// TIA Portal project "E95238_MCC1200_Sisecam_India" (V17) (continued)
TYPE "UDT_CapData_Tracking"
   STRUCT
      dTrackingHead : DInt;   // Tracking head on the circular buffer
      dTrackingTail : DInt;   // Tracking tail on the circular buffer
      dLastInsertIndex : DInt;   // Last insert index on circular
      dLastTargetLineValue_cmm : DInt;   // Last target line value [mm/100]
      dNextValidCapID : DInt;   // Next valid cap ID
      dLastValidCapID : DInt;   // Last valid cap ID
      dMutexCounter : DInt;   // Mutex counter for thread safe
      xInsertCapOnTrack : Bool;   // Insert cap on tracking
      timeLastAccessMutex : Time;   // Time of the last access mutex
      rgxNewCapAvailable : Array[0.."DMAXELEMWAKEUPNEWPLATE_IND"] of Bool;   // New cap available for other machines. Machines not used should be manually resetted
      tNewCapToInsert : "UDT_CapData";   // New cap to insert on tracking
      tLastPlacedCap : "UDT_CapData";   // Last placed cap on tracking
      rgtTrackCaps : Array[0.."DMAXTRACKCAP_IND"] of Struct   // Buffer of caps
         dEncValueHeadSnaproll_cmm : DInt;   // Encoder value on snap roll head [mm/100]
         dEncValueTailSnaproll_cmm : DInt;   // Encoder value on snap roll tail [mm/100]
         tCap : "UDT_CapData";   // Cap data
         rgxMachineExecMask : Array[0.."DMAXTRACKMACHINE_IND"] of Bool;   // Machine execution mask
      END_STRUCT;
      rgtTrackMachine : Array[0.."DMAXTRACKMACHINE_IND"] of Struct   // Tracking machine
         tUserData : Struct   // User data
            dSetDistanceSnap_cmm : DInt;   // Distance from snaproll [mm/100]
            dSetMachReacTime_ms : DInt;   // Machine reaction time [ms] (Positive to anticipate / Negative to delay)
            xGetPosReach : Bool;   // New cap arrive on position
            dGetUpstremIndex : DInt;   // Upstream cap position index
            dGetDownstreamIndex : DInt;   // Downstream cap position index
            dGetEncValueOnSnap_cmm : DInt;   // Encoder value on snaproll [mm/100]
         END_STRUCT;
         tAuxData : Struct   // Internal data for tracking
            dActualMachineEncValue_cmm : DInt;   // Actual machine encoder value [mm/100]
            dPrevCapIndex : DInt;   // Previous cap index
            dNextCapIndex : DInt;   // Next cap index
         END_STRUCT;
      END_STRUCT;
      tEmptyCap : "UDT_CapData";   // Cap with empty data (used for initialization)
      rgtTrackSearch : Array[0.."DMAXELEMTRACKSEARCH_IND"] of Struct   // Tracking search data
         xRequestSearchPlate : Bool;   // Request search plate
         xPlateFound : Bool;   // Plate found by tracking
         dRequestID : DInt;   // Number to identify the request
         dAnalyzedID : DInt;   // Number to identify the processed request
         dFoundTrackIndex : DInt;   // Plate pointer ID founded
         dSearchMode : DInt;   // Search mode (1=Limit head, 2=Limit tail 3=Both)
         dMinHeadPosition_cmm : DInt;   // Minimum head position distance from snaproll [mm/100]
         dMaxHeadPosition_cmm : DInt;   // Maximum head position distance from snaproll [mm/100]
         dMinTailPosition_cmm : DInt;   // Minumum tail position distance from snaproll [mm/100]
         dMaxTailPosition_cmm : DInt;   // Maximum tail position distance from snaproll [mm/100]
         tSearchRequest : Struct   // Search request
            xMainDestEqual : Bool;   // Main destination equal
            xLengthLessThan : Bool;   // Cap length is less than
            xCutDone : Bool;   // XCut is done
            xSpare_3 : Bool;
            xSpare_4 : Bool;
            xSpare_5 : Bool;
            xSpare_6 : Bool;
            xSpare_7 : Bool;
            xSpare_8 : Bool;
            xSpare_9 : Bool;
            xSpare_10 : Bool;
            xSpare_11 : Bool;
            xSpare_12 : Bool;
            xSpare_13 : Bool;
            xSpare_14 : Bool;
            xSpare_15 : Bool;
            xSpare_16 : Bool;
            xSpare_17 : Bool;
            xSpare_18 : Bool;
            xSpare_19 : Bool;
            xSpare_20 : Bool;
            xSpare_21 : Bool;
            xSpare_22 : Bool;
            xSpare_23 : Bool;
            xSpare_24 : Bool;
            xSpare_25 : Bool;
            xSpare_26 : Bool;
            xSpare_27 : Bool;
            xSpare_28 : Bool;
            xSpare_29 : Bool;
            xSpare_30 : Bool;
            xSpare_31 : Bool;
         END_STRUCT;
         tSearchData : Struct
            dMainDest_mask : LInt;   // Main destination mask
            dLength_cmm : DInt;   // Length [mm/100]
         END_STRUCT;
      END_STRUCT;
   END_STRUCT;
END_TYPE

// folder: 03_Encoder

TYPE "UDT_Encoder"
   STRUCT
      dActualEncoderCounter_cmm : DInt;   // Actual encoder counter [mm/100]
      rActSpeedValue_cmm_ms : Real;   // Actual speed value [(mm/100)/ms]
      dActSpeedValue_mm_min : DInt;   // Actual speed value [mm/min]
      rActSpeedValueFast_cmm_ms : Real;   // Actual speed value updated 500ms [(mm/100)/ms]
      dActSpeedValueFast_mm_min : DInt;   // Actual speed value updated 500ms [mm/min]
      dLastMeterValue_cmm : DInt;   // Last meter counter value [mm/100]
      dNextMeterValue_cmm : DInt;   // Next meter counter value [mm/100]
      rgxMetersForXcuts : Array[0.."DMAXXHEADS_IND"] of Bool;   // Meters signal for XCuts
      rgxMetersForYCuts : Array[0.."DMAXYCUTBRIDGE_IND"] of Bool;   // Meters signal for YCuts
      xMeterForMarkers : Bool;   // Meter signal for Markers
      xMeterForScanner : Bool;   // Meter signal for Scanner
   END_STRUCT;
END_TYPE

TYPE "LPD_typeCountFeedbackCh"
VERSION : 0.1
   STRUCT
      countValue : DInt := 16#0000;   // Current count value
      capturedValue : DInt := 16#0000;   // Last Capture value acquired
      measuredValue : Real := 0.0;   // Current measured value
      powerError : Bool := FALSE;   // Incorrect supply voltage L+
      encError : Bool := FALSE;   // Incorrect encoder signal
      ldError : Bool := FALSE;   // Error when loading via control interface
      reserved1 : Bool := FALSE;   // Reserved
      reserved2 : Bool := FALSE;   // Reserved
      reserved3 : Bool := FALSE;   // Reserved
      reserved4 : Bool := FALSE;   // Reserved
      reserved5 : Bool := FALSE;   // Reserved
      commActive : Bool := FALSE;   // Comm active
      resEventAck : Bool := FALSE;   // Reset of event bits active
      ldStsSlot0 : Bool := FALSE;   // Load request for Slot 0 detected and executed (toggling)
      ldStsSlot1 : Bool := FALSE;   // Load request for Slot 1 detected and executed (toggling)
      stsReady : Bool := FALSE;   // Digital on-board I/O started up and parameters assigned
      stsSwGate : Bool := FALSE;   // Software gate status
      reserved7 : Bool := FALSE;   // Reserved
      reserved8 : Bool := FALSE;   // Reserved
      stsDir : Bool := FALSE;   // Direction of last count value change
      stsCount : Bool := FALSE;   // Count pulse detected within last approx. 0.5 s
      stsGate : Bool := FALSE;   // Internal gate status
      stsDQ0 : Bool := FALSE;   // Status HSC DQ0
      stsDQ1 : Bool := FALSE;   // Status HSC DQ1
      stsDI0 : Bool := FALSE;   // Status HSC DI0
      stsDI1 : Bool := FALSE;   // Status HSC DI1
      stsDI2 : Bool := FALSE;   // Status HSC DI2
      eventZero : Bool := FALSE;   // Zero crossing has occurred
      eventUnderflow : Bool := FALSE;   // Underflow has occurred
      eventOverflow : Bool := FALSE;   // Overflow has occurred
      eventCompare0 : Bool := FALSE;   // Comparison event for DQ0 has occurred
      eventCompare1 : Bool := FALSE;   // Comparison event for DQ1 has occurred
      eventSync : Bool := FALSE;   // Synchronization has occurred
      eventCapture : Bool := FALSE;   // Capture event has occurred
      stsMeasInterval : Bool := FALSE;   // Count pulse detected in previous measuring interval
   END_STRUCT;
END_TYPE

TYPE "LPD_typeCountControlCh"
VERSION : 0.1
   STRUCT
      loadValue0 : DWord := 16#0000;   // Load value 0
      loadValue1 : DWord := 16#0000;   // Load value 1
      controlByte : Byte := B#16#00;   // Control byte load value
      swGate : Bool := FALSE;   // Software gate
      tmCtrlDQ0 : Bool := FALSE;   // Enable technological function DQ0
      tmCtrlDQ1 : Bool := FALSE;   // Enable technological function DQ1
      setDQ0 : Bool := FALSE;   // Set DQ0
      setDQ1 : Bool := FALSE;   // Set DQ1
      enSyncUp : Bool := FALSE;   // Enable upward synchronization
      enSyncDown : Bool := FALSE;   // Enable downward synchronization
      enCapture : Bool := FALSE;   // Enable capture function
      resError : Bool := FALSE;   // Reset of saved error states
      resEvent : Bool := FALSE;   // Reset of saved events
      reserved0 : Bool := FALSE;   // Reserved
      reserved1 : Bool := FALSE;   // Reserved
      reserved2 : Bool := FALSE;   // Reserved
      reserved3 : Bool := FALSE;   // Reserved
      reserved4 : Bool := FALSE;   // Reserved
      SetDir : Bool := FALSE;   // Count direction (with encoder without direction signal)
      reserved5 : Byte;   // Reserved
   END_STRUCT;
END_TYPE

// folder: 04_XCuts

TYPE "UDT_XCUT_DRIVE_INPUT"
   STRUCT
      rgxStatusBits : Struct
         xFault_EmergencyON : Bool := false;   // DN_SMAPP_FEMERGENCY_ON
         xFault_AuxPowerOFF : Bool := false;   // DN_SMAPP_FAUXPOWER_OFF
         xFault_InputPowerOFF : Bool := false;   // DN_SMAPP_FINPPOWER_OFF
         xFault_SafetyArea : Bool := false;   // DN_SMAPP_FSAFETYAREA
         xFault_Overtstroke : Bool := false;   // DN_SMAPP_FOVERSTROKE
         xFaultl_OverTemp : Bool := false;   // DN_SMAPP_FOVERTEMP
         xFault_CarriageNotDown : Bool := false;   // DN_SMAPP_FCARRIAGEDOWN
         xFault_MissingAir : Bool := false;   // DN_SMAPP_FMISSINGAIR
         xFault_AxisFault : Bool := false;   // DN_SMAPP_FAXISFAULT
         xFault_DriveNotEnable : Bool := false;   // DN_SMAPP_FDRIVENOENABLE
         xFault_TankOilEmpty : Bool := false;   // DN_SMAPP_FTANKOILEMPTY
         xFault_CarriageOff : Bool := false;   // DN_SMAPP_FCARRIAGEOFF
         xFault_ExtInpPower : Bool := false;   // DN_SMAPP_FEXTINPPOWER
         xFault_EmergencyLoc1 : Bool := false;   // DN_SMAPP_FLOCALEMERG_1
         xFault_EmergencyLoc2 : Bool := false;   // DN_SMAPP_FLOCALEMERG_2
         xFault_EmergencyLoc3 : Bool := false;   // DN_SMAPP_FLOCALEMERG_3
         xStatus_AxisOnline : Bool := false;   // DN_SMAPP_AXISONLINE
         xStatus_AxisReady : Bool := false;   // DN_SMAPP_AXISREADY
         xStatus_HomeProgress : Bool := false;   // DN_SMAPP_HOMEPROGRESS
         xStatus_MoveProgress : Bool := false;   // DN_SMAPP_MOVEPROGRESS
         xStatus_MoveProgrNick : Bool := false;   // DN_SMAPP_MOVEPROGRESSNICK
         xStatus_InvertReady : Bool := false;   // DN_SMAPP_INVERTERREADY
         xStatus_BridgeEnabled : Bool := false;   // DN_SMAPP_BRIDGEENABLED
         xStatus_AxisSyncronized : Bool := false;   // DN_SMAPP_AXISSYNCRONIZED
         xStatus_ButtonEnabled : Bool;   // Button enabled
         xStatus_xSpare17 : Bool;   // Spare
         xStatus_xSpare18 : Bool;   // Spare
         xStatus_xSpare19 : Bool;   // Spare
         xStatus_xSpare20 : Bool;   // Spare
         xStatus_xSpare21 : Bool;   // Spare
         xStatus_xSpare22 : Bool;   // Spare
         xStatus_xSpare23 : Bool;   // Spare
      END_STRUCT;
      dCarriagePos_dmm : DInt := 0;   // DN_SMAPP_CARRIAGEPOS [mm/10]
      dLehrPosition_cmm : DInt := 0;   // DN_SMAPP_LEHRPOSITION [mm/100]
      dLehrSpeed_cmm_min : DInt := 0;   // DN_SMAPP_LEHRSPEED [mm/10/min]
      dErrorCode : DInt := 0;   // DN_SMAPP_ERRORCODE
      dMissionDone : DInt := 0;   // DN_SMAPP_MISSIONDONE
      dMissionUnDone : DInt := 0;   // DN_SMAPP_MISSION_UNDONE
      iLiveCounter : Int := 0;   // DN_SMAPP_LIVECOUNTER
      iTimeHeadDown_ms : Int;   // Time head down% [ms]
   END_STRUCT;
END_TYPE

TYPE "UDT_XCUT_DRIVE_OUTPUT"
   STRUCT
      rgxControlBits : Struct
         xSpare0 : Bool;
         xSpare1 : Bool;
         xSpare2 : Bool;
         xSpare3 : Bool;
         xFaultReset : Bool := false;   // DN_PLC_FAULTRESET
         xEnableBridge : Bool := false;   // DN_PLC_ENABLEBRIDGE
         xDisableBridge : Bool := false;   // DN_PLC_DISABLEBRIDGE
         xSimulationMode : Bool := false;   // DN_PLC_SIMULATIONMODE
         xDisableRequest : Bool;   // DN_PLC_DISABLEREQUEST
         xSpare9 : Bool;
         xSpare10 : Bool;
         xSpare11 : Bool;
         xSpare12 : Bool;
         xSpare13 : Bool;
         xSpare14 : Bool;
         xSpare15 : Bool;
         xSpare16 : Bool;
         xSpare17 : Bool;
         xSpare18 : Bool;
         xSpare19 : Bool;
         xSpare20 : Bool := false;
         xSpare21 : Bool := false;
         xSpare22 : Bool := false;
         xSpare23 : Bool := false;
         xSpare24 : Bool;
         xSpare25 : Bool;
         xSpare26 : Bool;
         xSpare27 : Bool;
         xSpare28 : Bool;
         xSpare29 : Bool;
         xSpare30 : Bool;
         xSpare31 : Bool;
      END_STRUCT;
      dBridgeAngle_degre_10000 : DInt := 0;   // DN_PLC_BRIDGEANGLE
      dHeadDownPos_dmm : DInt := 0;   // DN_PLC_HEADDOWNPOS
      dHeadRisePos_dmm : DInt := 0;   // DN_PLC_HEADRISEPOS
      iReturnSpeed_rpm : Int := 0;   // DN_PLC_RETURNSPEED
      iTimeHeadDown_ms : Int := 0;   // DN_PLC_TIMEHEADDOWN
      iTimeHeadUp_ms : Int := 0;   // DN_PLC_TIMEHEADUP
      iLubAdvanceTime_ms : Int := 0;   // DN_PLC_LUBADVANCETIME
      iLubDelayTime_ms : Int := 0;   // DN_PLC_LUBDELAYTIME
      iTimeHeadAct_ms : Int := 0;   // DN_PLC_TIMEHEADACTIV
      iTimeHeadDeactiv_ms : Int := 0;   // DN_PLC_TIMEHEADDEACTIV
      dPressure_mN : DInt := 0;   // DN_PLC_PRESSURE
      dMissionID : DInt := 0;   // DN_PLC_MISSIONID
      dMissionCounter : DInt := 0;   // DN_PLC_MISSIONCOUNTER
      dSyncroCounter : DInt := 0;   // DN_PLC_SYNCROCOUNTER
      iLiveCounter : Int := 0;   // DN_PLC_LIVECOUNTER
   END_STRUCT;
END_TYPE

TYPE "UDT_XCUT_AXIS_REF"
   STRUCT
      udi_ModbusAddress_read : UDInt;
      di_ParameterReadValue : DInt;
      x_CommandReadParameter : Bool;
      x_StatusReadParameter_OK : Bool;
      x_StatusReadParameter_Error : Bool;
      udi_ModbusAddress_write : UDInt;
      di_ParameterWriteValue : DInt;
      x_CommandWriteParameter : Bool;
      x_Status_WriteParameter_OK : Bool;
      x_Status_WriteParameter_Error : Bool;
   END_STRUCT;
END_TYPE

// folder: 05_YCuts

TYPE "UDT_YCut_IdeviceToBridge"
   STRUCT
      dSpare1 : Array[0..2] of DInt;
      xCycleON : Bool;
      xResetAnomaly : Bool;
      xResetBuffers : Bool;
      xGlassBreak : Bool;
      xPLCActive0 : Bool;
      xPLCActive1 : Bool;
      xQLTplate : Bool;
      xSpare2 : Bool;
      xSpare3 : Bool;
      xSpare4 : Bool;
      xSpare5 : Bool;
      xSpare6 : Bool;
      xSpare7 : Bool;
      xSpare8 : Bool;
      xSpare9 : Bool;
      xSpare10 : Bool;
      xStatusSpare : Array[0..15] of Bool;
      dSpare2 : Array[0..7] of DInt;
      iSpare : Int;
   END_STRUCT;
END_TYPE

TYPE "UDT_YCut_IdeviceFromBridge"
   STRUCT
      dProcessingIDPlate : DInt;   // Processing ID Plate [Num]
      dSpare1 : DInt;
      dBridgeStatus : DInt;
      rgxStatus : Array[0..31] of Bool;   // Status heads
      rgdHeadsPositions_cmm : Array[0..15] of DInt;   // Head #x position status
      rgxHeadStatus : Array[0..15] of Bool;   // Head #x enabled
      rgxCuttingStatus : Array[0..15] of Bool;   // Head #x cuuting status
      rgdHeadsPressure : Array[0..15] of DInt;   // Head #x Pressure [mN]
      rgrHeadsSpace : Array[0..15] of Real;   // Head #x Distance [Km]
      iFireOffset_ON : Int;   // All head fire on offset
      iFireOffset_OFF : Int;   // All head fire off offset
      iSpare : Int;
      dSpare : Array[0..7] of DInt;
   END_STRUCT;
   // // rgxStatus[0] : Glass break in progress
   // // rgxStatus[1] : Liftup pushbutton engaged
   // // rgxStatus[2] : Bridge enabled
   // // rgxStatus[3] : Bridge locked
   // // rgxStatus[8] : Fire offset calibration
   // // rgxStatus[4] : Status heads
   // // rgxStatus[5] : Status heads
   // // rgxStatus[6] : Status heads
   // // rgxStatus[7] : Status heads
   // // rgxStatus[9] : Status heads
   // // rgxStatus[10] : Status heads
   // // rgxStatus[11] : Status heads
   // // rgxStatus[12] : Status heads
   // // rgxStatus[13] : Status heads
   // // rgxStatus[14] : Status heads
   // // rgxStatus[15] : Status heads
   // // rgxStatus[16] : Status heads
   // // rgxStatus[17] : Status heads
   // // rgxStatus[18] : Status heads
   // // rgxStatus[19] : Status heads
   // // rgxStatus[20] : Status heads
   // // rgxStatus[21] : Status heads
   // // rgxStatus[22] : Status heads
   // // rgxStatus[23] : Status heads
   // // rgxStatus[24] : Status heads
   // // rgxStatus[25] : Status heads
   // // rgxStatus[26] : Status heads
   // // rgxStatus[27] : Status heads
   // // rgxStatus[28] : Status heads
   // // rgxStatus[29] : Status heads
   // // rgxStatus[30] : Status heads
   // // rgxStatus[31] : Status heads
END_TYPE

// folder: 06_Markers

TYPE "UDT_Marker_Mission_Data"
   STRUCT
      dPlateID : DInt;   // Defect plate ID
      dMissionID : DInt;   // Mission ID
      dMarkerID : DInt;   // Marker ID (0=Auto, 1=M#1, 2=M#2, 3=M#3, 4=M#4)
      dXPosition_cmm : DInt;   // Marker counter X position [mm/100]
      dYPosition_cmm : DInt;   // Marker Y position [mm/100]
      dSpotSpace_cmm : DInt;   // Spot space [mm/100]
   END_STRUCT;
END_TYPE

TYPE "UDT_Marker_IDeviceToBridge"
   STRUCT
      xCycleON : Bool;   // Cycle ON
      xResetAnomaly : Bool;   // Reset anomaly
      xResetBuffers : Bool;   // Reset buffer
      xGlassBreak : Bool;   // Glass break under the bridge
      Spare_x4 : Bool;
      Spare_x5 : Bool;
      Spare_x6 : Bool;
      Spare_x7 : Bool;
      Spare_x8 : Bool;
      Spare_x9 : Bool;
      Spare_x10 : Bool;
      Spare_x11 : Bool;
      Spare_x12 : Bool;
      Spare_x13 : Bool;
      Spare_x14 : Bool;
      Spare_x15 : Bool;
      xStatusSpare : Array[0..15] of Bool;
      dSpare2 : Array[0..7] of DInt;
   END_STRUCT;
END_TYPE

TYPE "UDT_Marker_IDeviceFromBridge"
   STRUCT
      rgdHeadsPositions_cmm : Array[0.."DMAXMARKERS_IND"] of DInt;   // Head #x position status
      rgdBridgeProdModeActual : Array[0.."DMAXMARKERS_IND"] of DInt;   // Production modality actual (1=Out of production 3=In production 8=Out of production request 9=In production request)
      rgdDistanceFromSnaproll_cmm : Array[0.."DMAXMARKERS_IND"] of DInt;   // Distance from snaproll [mm/100]
      rgdDistanceFromCenterLine_cmm : Array[0.."DMAXMARKERS_IND"] of DInt;   // Distance from center line [mm/100]
      rgdSpraySpace_cmm : Array[0.."DMAXMARKERS_IND"] of DInt;   // Markers spray time [ms]
      dSpare : Array[0..4] of DInt;
   END_STRUCT;
END_TYPE

// folder: 07_Z300

TYPE "UDT_iDeviceZ301--->Z200"
   STRUCT
      Z300 : Struct
         tAuxBits : Struct   // Auxiliary bits
            xCleaningActiveHL : Bool;   // Cleaning active lamp
            xLineOK : Bool;   // Line is ok
            xZ301AnomalyHL : Bool;   // Z301 anomaly lamp
            xZ302AnomalyHL : Bool;   // Z302 anomaly lamp
            xCPUAActive : Bool;   // CPU A is active
            xCPUBActive : Bool;   // CPU B is active
            xThicknessChangeActive : Bool;   // Thickness change modality is active
            xSpare10 : Bool;
            xSpare11 : Bool;
            xSpare12 : Bool;
            xSpare13 : Bool;
            xSpare14 : Bool;
            xSpare15 : Bool;
            xSpare22 : Bool;
            xSpare23 : Bool;
            xSpare24 : Bool;
            xSpare25 : Bool;
            xSpare26 : Bool;
            xSpare27 : Bool;
            xSpare28 : Bool;
            xSpare29 : Bool;
            xSpare30 : Bool;
            xSpare31 : Bool;
         END_STRUCT;
         tCulletSystem : Struct
            xHoldBreakerT2 : Bool;
            xSpare1 : Bool;
            xSpare2 : Bool;
            xSpare3 : Bool;
            xSpare4 : Bool;
            xSpare5 : Bool;
            xSpare6 : Bool;
            xSpare7 : Bool;
            xSpare8 : Bool;
            xSpare9 : Bool;
            xSpare10 : Bool;
            xSpare11 : Bool;
            xSpare12 : Bool;
            xSpare13 : Bool;
            xSpare14 : Bool;
            xSpare15 : Bool;
            xSpare16 : Bool;
            xSpare17 : Bool;
            xSpare18 : Bool;
            xSpare19 : Bool;
            xSpare20 : Bool;
            xSpare21 : Bool;
            xSpare22 : Bool;
            xSpare23 : Bool;
            xSpare24 : Bool;
            xSpare25 : Bool;
            xSpare26 : Bool;
            xSpare27 : Bool;
            xSpare28 : Bool;
            xSpare29 : Bool;
            xSpare30 : Bool;
            xSpare31 : Bool;
         END_STRUCT;
         dLineSpeed_mm_min : DInt;   // Line speed [mm/min]
         dSpeedZone1_mm_min : DInt;   // Speed zone 1 acceleration [mm/min]
         dDownstreamSpeedContrast_mm_min : DInt;
         rgdSpare : Array[0..4] of DInt;
      END_STRUCT;
      Z200 : Struct
         dLherSpeed_Enc1 : DInt;   // Lher Speed Encoder 1 pulse
         dLherSpeed_Enc2 : DInt;   // Lher Speed Encoder 2 pulse
         IN_MCC1201 : Struct
            "xA.E20.0" : Bool;
            "xA.E20.1" : Bool;
            "xA.E20.2" : Bool;
            "xA.E20.3" : Bool;
            "xA.E20.4" : Bool;
            "xA.E20.5" : Bool;
            "xA.E20.6" : Bool;
            "xA.E20.7" : Bool;
            "xA.E21.0" : Bool;
            "xA.E21.1" : Bool;
            "xA.E21.2" : Bool;
            "xA.E21.3" : Bool;
            "xA.E21.4" : Bool;
            "xA.E21.5" : Bool;
            "xA.E21.6" : Bool;
            "xA.E21.7" : Bool;
            "xA.E80.0" : Bool;
            "xA.E80.1" : Bool;
            "xA.E80.2" : Bool;
            "xA.E80.3" : Bool;
            "xA.E80.4" : Bool;
            "xA.E80.5" : Bool;
            "xA.E80.6" : Bool;
            "xA.E80.7" : Bool;
            "xA.E81.0" : Bool;
            "xA.E81.1" : Bool;
            "xA.E81.2" : Bool;
            "xA.E81.3" : Bool;
            "xA.E81.4" : Bool;
            "xA.E81.5" : Bool;
            "xA.E81.6" : Bool;
            "xA.E81.7" : Bool;
            "xA.E82.0" : Bool;
            "xA.E82.1" : Bool;
            "xA.E82.2" : Bool;
            "xA.E82.3" : Bool;
            "xA.E82.4" : Bool;
            "xA.E82.5" : Bool;
            "xA.E82.6" : Bool;
            "xA.E82.7" : Bool;
            "xA.E83.0" : Bool;
            "xA.E83.1" : Bool;
            "xA.E83.2" : Bool;
            "xA.E83.3" : Bool;
            "xA.E83.4" : Bool;
            "xA.E83.5" : Bool;
            "xA.E83.6" : Bool;
            "xA.E83.7" : Bool;
            "xA.E32.0" : Bool;   // PhotoM202
            "xA.E32.1" : Bool;   // PhotoM202
            "xA.E32.2" : Bool;   // PhotoM202
            "xA.E32.3" : Bool;   // PhotoM202
            "xA.E32.4" : Bool;   // PhotoM202
            "xA.E32.5" : Bool;   // PhotoM202
            "xA.E32.6" : Bool;   // PhotoM202
            "xA.E32.7" : Bool;   // PhotoM202
            "xA.E33.0" : Bool;   // PhotoM202
            "xA.E33.1" : Bool;   // PhotoM202
            "xA.E33.2" : Bool;
            "xA.E33.3" : Bool;
            "xA.E33.4" : Bool;
            "xA.E33.5" : Bool;
            "xA.E33.6" : Bool;
            "xA.E33.7" : Bool;
            "xA.E34.0" : Bool;
            "xA.E34.1" : Bool;
            "xA.E34.2" : Bool;
            "xA.E34.3" : Bool;
            "xA.E34.4" : Bool;
            "xA.E34.5" : Bool;
            "xA.E34.6" : Bool;
            "xA.E34.7" : Bool;
            "xA.E35.0" : Bool;
            "xA.E35.1" : Bool;
            "xA.E35.2" : Bool;
            "xA.E35.3" : Bool;
            "xA.E35.4" : Bool;
            "xA.E35.5" : Bool;
            "xA.E35.6" : Bool;
            "xA.E35.7" : Bool;
            "xA.E36.0" : Bool;
            "xA.E36.1" : Bool;
            "xA.E36.2" : Bool;
            "xA.E36.3" : Bool;
            "xA.E36.4" : Bool;
            "xA.E36.5" : Bool;
            "xA.E36.6" : Bool;
            "xA.E36.7" : Bool;
            "xA.E37.0" : Bool;
            "xA.E37.1" : Bool;
            "xA.E37.2" : Bool;
            "xA.E37.3" : Bool;
            "xA.E37.4" : Bool;
            "xA.E37.5" : Bool;
            "xA.E37.6" : Bool;
            "xA.E37.7" : Bool;
            "xA.E38.0" : Bool;
            "xA.E38.1" : Bool;
            "xA.E38.2" : Bool;
            "xA.E38.3" : Bool;
            "xA.E38.4" : Bool;
            "xA.E38.5" : Bool;
            "xA.E38.6" : Bool;
            "xA.E38.7" : Bool;
            "xA.E39.0" : Bool;
            "xA.E39.1" : Bool;
            "xA.E39.2" : Bool;
            "xA.E39.3" : Bool;
            "xA.E39.4" : Bool;
            "xA.E39.5" : Bool;
            "xA.E39.6" : Bool;
            "xA.E39.7" : Bool;
            rtgSpare : Array[0..9] of Int;
         END_STRUCT;
         IN_MCC1301 : Struct
            "xE.E108.0" : Bool;
            "xE.E108.1" : Bool;
            "xE.E108.2" : Bool;
            "xE.E108.3" : Bool;
            "xE.E108.4" : Bool;
            "xE.E108.5" : Bool;
            "xE.E108.6" : Bool;
            "xE.E108.7" : Bool;
            xSpare8 : Bool;
            xSpare9 : Bool;
            xSpare10 : Bool;
            xSpare11 : Bool;
            xSpare12 : Bool;
            xSpare13 : Bool;
            xSpare14 : Bool;
            xSpare15 : Bool;
            xSpare22 : Bool;
            xSpare23 : Bool;
            xSpare24 : Bool;
            xSpare25 : Bool;
            xSpare26 : Bool;
            xSpare27 : Bool;
            xSpare28 : Bool;
            xSpare29 : Bool;
            xSpare30 : Bool;
            xSpare31 : Bool;
         END_STRUCT;
         rtgSpare : Array[0..6] of Int;
      END_STRUCT;
   END_STRUCT;
END_TYPE

TYPE "UDT_iDeviceZ301<---Z200"
   STRUCT
      Z300 : "UDT_iDeviceZ301<---Z200_INO";
      MCC_Out : "UDT_iDevice_MCC1201<---Mcc1200_OUT";
   END_STRUCT;
END_TYPE

TYPE "UDT_iDeviceZ301<---Z200_INO"
   STRUCT
      Z300 : Struct
         tCulletSystem : Struct
            xBreakerT2Ready : Bool;
            xSpare1 : Bool;
            xSpare2 : Bool;
            xSpare3 : Bool;
            xSpare4 : Bool;
            xSpare5 : Bool;
            xSpare6 : Bool;
            xSpare7 : Bool;
            xSpare8 : Bool;
            xSpare9 : Bool;
            xSpare10 : Bool;
            xSpare11 : Bool;
            xSpare12 : Bool;
            xSpare13 : Bool;
            xSpare14 : Bool;
            xSpare15 : Bool;
            xSpare16 : Bool;
            xSpare17 : Bool;
            xSpare18 : Bool;
            xSpare19 : Bool;
            xSpare20 : Bool;
            xSpare21 : Bool;
            xSpare22 : Bool;
            xSpare23 : Bool;
            xSpare24 : Bool;
            xSpare25 : Bool;
            xSpare26 : Bool;
            xSpare27 : Bool;
            xSpare28 : Bool;
            xSpare29 : Bool;
            xSpare30 : Bool;
            xSpare31 : Bool;
         END_STRUCT;
      END_STRUCT;
   END_STRUCT;
END_TYPE

TYPE "UDT_iDevice_MCC1201<---Mcc1200_OUT"
   STRUCT
      Z200 : Struct
         tOUT_Mcc1201 : Struct
            "xA86.0" : Bool;
            "xA86.1" : Bool := false;
            "xA86.2" : Bool := false;
            "xA86.3" : Bool := false;
            "xA86.4" : Bool := false;
            "xA86.5" : Bool := false;
            "xA86.6" : Bool := false;
            "xA86.7" : Bool := false;
            "xA87.0" : Bool := false;
            "xA87.1" : Bool := false;
            "xA87.2" : Bool := false;
            "xA87.3" : Bool := false;
            "xA87.4" : Bool := false;
            "xA87.5" : Bool := false;
            "xA87.6" : Bool := false;
            "xA87.7" : Bool := false;
            "xA44.0" : Bool := false;
            "xA44.1" : Bool := false;
            "xA44.2" : Bool := false;
            "xA44.3" : Bool := false;
            "xA44.4" : Bool := false;
            "xA44.5" : Bool := false;
            "xA44.6" : Bool := false;
            "xA44.7" : Bool := false;
            "xA45.0" : Bool := false;
            "xA45.1" : Bool := false;
            "xA45.2" : Bool := false;
            "xA45.3" : Bool := false;
            "xA45.4" : Bool := false;
            "xA45.5" : Bool := false;
            "xA45.6" : Bool := false;
            "xA45.7" : Bool := false;
            "xA46.0" : Bool := false;
            "xA46.1" : Bool := false;
            "xA46.2" : Bool := false;
            "xA46.3" : Bool := false;
            "xA46.4" : Bool := false;
            "xA46.5" : Bool := false;
            "xA46.6" : Bool := false;
            "xA46.7" : Bool := false;
            "xA47.0" : Bool := false;
            "xA47.1" : Bool := false;
            "xA47.2" : Bool := false;
            "xA47.3" : Bool := false;
            "xA47.4" : Bool := false;
            "xA47.5" : Bool := false;
            "xA47.6" : Bool := false;
            "xA47.7" : Bool := false;
         END_STRUCT;
         rgdSpare_0 : Array[0..4] of DInt;
         tOUT_Mcc1301 : Struct
            "xE.A126.0" : Bool;
            "xE.A126.1" : Bool;
            "xE.A126.2" : Bool;
            "xE.A126.3" : Bool;
            "xE.A126.4" : Bool;
            "xE.A126.5" : Bool;
            "xE.A126.6" : Bool;
            "xE.A126.7" : Bool;
            xSpare8 : Bool;
            xSpare9 : Bool;
            xSpare10 : Bool;
            xSpare11 : Bool;
            xSpare12 : Bool;
            xSpare13 : Bool;
            xSpare14 : Bool;
            xSpare15 : Bool;
            xSpare16 : Bool;
            xSpare17 : Bool;
            xSpare18 : Bool;
            xSpare19 : Bool;
            xSpare20 : Bool;
            xSpare21 : Bool;
            xSpare22 : Bool;
            xSpare23 : Bool;
            xSpare24 : Bool;
            xSpare25 : Bool;
            xSpare26 : Bool;
            xSpare27 : Bool;
            xSpare28 : Bool;
            xSpare29 : Bool;
            xSpare30 : Bool;
            xSpare31 : Bool;
         END_STRUCT;
         rgdSpare_1 : Array[0..4] of DInt;
      END_STRUCT;
      Z300 : Struct
         tAuxBits : Struct
            xGlassBreakOut : Bool;   // Glass breakout
            xEmptyingLineArea301 : Bool;   // Not used Emptying lire area 301
            xResetAnomaly301 : Bool;   // Not used Reset anomaly 301
            xResetAnomaly302 : Bool;   // Not used Reset anomaly 302
            xCycleOn : Bool;   // Cycle ON
            xSirenCulletStop : Bool;   // Not used Siren cullet stop
            xStartCycleRequest : Bool;   // Not used Start cycle request
            xBypassGlassLengthCheck : Bool;   // Not used Bypass glass length check due stripe
            xCPUAActive : Bool;   // CPU A Active
            xCPUBActive : Bool;   // CPU B Active
            xStopEmptyingLineArea301 : Bool;   // Not used Stop emptying line area 301
            xSpare11 : Bool;
            xSpare12 : Bool;
            xSpare13 : Bool;
            xSpare14 : Bool;
            xSpare15 : Bool;
            xBreakOUTDoneCheck : Bool;
            xSelectionDriveA : Bool;
            xSelectionDriveB : Bool;
            xSpare19 : Bool;
            xSpare20 : Bool;
            xSpare21 : Bool;
            xSpare22 : Bool;
            xSpare23 : Bool;
            xSpare24 : Bool;
            xSpare25 : Bool;
            xSpare26 : Bool;
            xSpare27 : Bool;
            xSpare28 : Bool;
            xSpare29 : Bool;
            xSpare30 : Bool;
            xSpare31 : Bool;
         END_STRUCT;
         dLehrSpeed_to_Conv_mm_min : DInt;   // Lehr speed [mm/min]
         dDownstremConstrastPosition_cmm : DInt;   // Downstream constrast position [mm/100] (0 is snaproll)
         iSpare : Int;
         rgdSpare : Array[0..7] of DInt;
      END_STRUCT;
   END_STRUCT;
END_TYPE

TYPE "UDT_CapData_Z300"
   STRUCT
      dID : DInt;   // Cap ID [Num]
      dProductionID : DInt;   // Cap production ID
      dLength_cmm : DInt;   // Cap length [mm/100]
      dWidth_cmm : DInt;   // Cap total width [mm/100]
      dThick_cmm : DInt;   // Cap thickness [mm/100]
      dGap_cmm : DInt;   // Cap Gap [mm/100]
      dIndex : DInt;   // Cap index number in convoy [Num] (0=First cap in convoy)
      dFormat : DInt;   // Plate format [Num] (1=JS 2=Les 3=SSS)
      dNumLites : DInt;   // Number of lites in cap [Num]
      dReqGapForConv_cmm : DInt;   // Request gap beetween caps for convoy creation [mm/100]
      dMaxCapInConv : DInt;   // Maximum number of cap in convoy
      dConvTotLength_cmm : DInt;   // Total length of the convoy [mm/100]
      dMinWidth_cmm : DInt;   // Shortest width in use [mm/100]
      dMaxWidth_cmm : DInt;   // Biggest width in use [mm/100]
      dGrossWidth_cmm : DInt;   // Cap gross width [mm/100]
      dNetWidth_cmm : DInt;   // Cap net width [mm/100]
      dDEdgeOpSide_cmm : DInt;   // Double edge dimension - operator side [mm/100]
      dDEdgeOppOpSide_cmm : DInt;   // Double edge dimension - opposite operator side [mm/100]
      dTEdgeOpSide_cmm : DInt;   // Triple edge dimension - operator side [mm/100]
      dTEdgeOppOpSide_cmm : DInt;   // Triple edge dimension - opposite operator side [mm/100]
      dCutWander_cmm : DInt;   // Cap cut wander (- Op. Side + Oppo. Op. Side) [mm/100]
      dStackerModality : DInt;   // Staker Modality (0:MonoPortrate , 1: MonoLandascape , 10:SteroPortrate , 11: SteroLandascape)
      dStackerMode : DInt;   // Staker Mode (0: Air , 1: TIN)
      dColor : DInt;   // Color code [Num]
      xFixedCapProduction : Bool;   // Fixed cap production
      strColorDescr : String["DSTRSIZEDESCR"];   // Color description [Text]
      tFlagTrim : Struct
         xByYCut1 : Bool;
         xByYCut2 : Bool;
         xTrim3OpSide : Bool;
         xTrim2OpSide : Bool;
         xTrim1OpSide : Bool;
         xTrim1OppOpSide : Bool;
         xTrim2OppOpSide : Bool;
         xTrim3OppOpSide : Bool;
         rgxIntCut : Array[0..15] of Bool;
         xOptSelvedgeSel : Bool;
         xOptSplitBarSel : Bool;
         xOptSepRollSel : Bool;
         tSelvedge : Struct
            dRequestTrim3OpSide : DInt;
            dRequestTrim2OpSide : DInt;
            dRequestTrim1OpSide : DInt;
            dRequestTrim3OppOpSide : DInt;
            dRequestTrim2OppOpSide : DInt;
            dRequestTrim1OppOpSide : DInt;
            dDoneTrim3OpSide : DInt;
            dDoneTrim2OpSide : DInt;
            dDoneTrim1OpSide : DInt;
            dDoneTrim3OppOpSide : DInt;
            dDoneTrim2OppOpSide : DInt;
            dDoneTrim1OppOpSide : DInt;
         END_STRUCT;
         tSplitBar : Array[0..15] of Struct
            dRequestSnapCut : DInt;
            dDoneSnapCut : DInt;
         END_STRUCT;
         tSepRoll : Array[0..15] of Struct
            rgxRequestSeparator : Array[0..15] of Bool;
            rgxDoneSeparator : Array[0..15] of Bool;
         END_STRUCT;
         rgxXCutDoneHead : Array[0..15] of Bool;
         rgxXCutDoneTail : Array[0..15] of Bool;
         rgxYCutHeadDone : Array[0..15] of Bool;
      END_STRUCT;
      tRequests : Struct   // Lavoration request on cap
         Spare1 : Bool;
         Spare2 : Bool;
         Spare3 : Bool;
         Spare4 : Bool;
         Spare5 : Bool;
         Spare6 : Bool;
         Spare7 : Bool;
         Spare8 : Bool;
         Spare9 : Bool;
         Spare10 : Bool;
         Spare11 : Bool;
         Spare12 : Bool;
         Spare13 : Bool;
         Spare14 : Bool;
         Spare15 : Bool;
         Spare16 : Bool;
         Spare17 : Bool;
         Spare18 : Bool;
         Spare19 : Bool;
         Spare20 : Bool;
         Spare21 : Bool;
         Spare22 : Bool;
         Spare23 : Bool;
         Spare24 : Bool;
         Spare25 : Bool;
         Spare26 : Bool;
         Spare27 : Bool;
         Spare28 : Bool;
         Spare29 : Bool;
         Spare30 : Bool;
         Spare31 : Bool;
         Spare32 : Bool;
      END_STRUCT;
      tDone : Struct   // Lavoration done on cap
         Spare1 : Bool;
         Spare2 : Bool;
         Spare3 : Bool;
         Spare4 : Bool;
         Spare5 : Bool;
         Spare6 : Bool;
         Spare7 : Bool;
         Spare8 : Bool;
         Spare9 : Bool;
         Spare10 : Bool;
         Spare11 : Bool;
         Spare12 : Bool;
         Spare13 : Bool;
         Spare14 : Bool;
         Spare15 : Bool;
         Spare16 : Bool;
         Spare17 : Bool;
         Spare18 : Bool;
         Spare19 : Bool;
         Spare20 : Bool;
         Spare21 : Bool;
         Spare22 : Bool;
         Spare23 : Bool;
         Spare24 : Bool;
         Spare25 : Bool;
         Spare26 : Bool;
         Spare27 : Bool;
         Spare28 : Bool;
         Spare29 : Bool;
         Spare30 : Bool;
         Spare31 : Bool;
         Spare32 : Bool;
      END_STRUCT;
      rgtLites : Array[0..12] of Struct   // Lites data
         dID : DInt;   // Lite ID [Num]
         dProductionID : DInt;   // Production ID [Num]
         strProdDescr : String["DSTRSIZEDESCR"];   // Production description [Text]
         dQualityID : DInt;   // Quality ID [Num]
         strQualityDescr : String["DSTRSIZEDESCR"];   // Quality description [Text]
         dCameraRecipeID : DInt;   // Camera recipe ID [Num]
         dWidth_cmm : DInt;   // Width [mm/100]
         dBarycentre_cmm : DInt;   // Barycentre [mm/100]
         dCulletCause_cmm : DInt;   // Cullet cause [mm/100]
         rgxLayers : Array[0.."DMAXPROTLAYER_IND"] of Bool;   // Protection layers requested
         rgxOrigin : Array[0.."DNUMBEROFDESTINATION_Z300"] of Bool;
         rgxMain : Array[0.."DNUMBEROFDESTINATION_Z300"] of Bool;
         rgxAlternative : Array[0.."DNUMBEROFDESTINATION_Z300"] of Bool;
         rgx2ndDestination : Array[0.."DNUMBEROFDESTINATION_Z300"] of Bool;
         tRequests : Struct   // Request for lites
            xReqGeoIspection : Bool;
            xReqPowderA : Bool;
            xReqPowderB : Bool;
            Spare4 : Bool;
            Spare5 : Bool;
            Spare6 : Bool;
            Spare7 : Bool;
            Spare8 : Bool;
            Spare9 : Bool;
            Spare10 : Bool;
            Spare11 : Bool;
            Spare12 : Bool;
            Spare13 : Bool;
            Spare14 : Bool;
            Spare15 : Bool;
            Spare16 : Bool;
            Spare17 : Bool;
            Spare18 : Bool;
            Spare19 : Bool;
            Spare20 : Bool;
            Spare21 : Bool;
            Spare22 : Bool;
            Spare23 : Bool;
            Spare24 : Bool;
            Spare25 : Bool;
            Spare26 : Bool;
            Spare27 : Bool;
            Spare28 : Bool;
            Spare29 : Bool;
            Spare30 : Bool;
            Spare31 : Bool;
            Spare32 : Bool;
         END_STRUCT;
         tDone : Struct   // Done for lites
            Spare1 : Bool;
            Spare2 : Bool;
            Spare3 : Bool;
            Spare4 : Bool;
            Spare5 : Bool;
            Spare6 : Bool;
            Spare7 : Bool;
            Spare8 : Bool;
            Spare9 : Bool;
            Spare10 : Bool;
            Spare11 : Bool;
            Spare12 : Bool;
            Spare13 : Bool;
            Spare14 : Bool;
            Spare15 : Bool;
            Spare16 : Bool;
            Spare17 : Bool;
            Spare18 : Bool;
            Spare19 : Bool;
            Spare20 : Bool;
            Spare21 : Bool;
            Spare22 : Bool;
            Spare23 : Bool;
            Spare24 : Bool;
            Spare25 : Bool;
            Spare26 : Bool;
            Spare27 : Bool;
            Spare28 : Bool;
            Spare29 : Bool;
            Spare30 : Bool;
            Spare31 : Bool;
            Spare32 : Bool;
         END_STRUCT;
         xSaturationPlate : Bool;
      END_STRUCT;
   END_STRUCT;
END_TYPE

// folder: 08_Report

TYPE "UDT_RP_MessageContMerge_v2"
VERSION : 0.1
   STRUCT
      xInitialized : Bool;   // The block is correctly initialized
      dNumOfMessage : DInt;   // Actual number of messages in buffer
      dMaxNumOfMessage : DInt;   // Maximum number of message in buffer
      rgtMessages : Array[0..12] of "UDT_RP_Message_v2";   // Array of messages
   END_STRUCT;
END_TYPE

TYPE "UDT_RP_TankMessages"
   STRUCT
      dNumberOfMessage : DInt;   // Number of message on tank
      rgtMessages : Array[0.."DMAXNUMMESSAGETANK_IND"] of "UDT_RP_Message_v2";
   END_STRUCT;
END_TYPE

TYPE "UDT_RP_AddMessageCont_v2"
VERSION : 0.1
   STRUCT
      xInitialized : Bool;   // The block is correctly initialized
      dNumOfMessage : DInt;   // Actual number of messages in buffer
      dMaxNumOfMessage : DInt;   // Maximum number of message in buffer
      rgtMessages : Array[0..99] of "UDT_RP_Message_v2";   // Array of messages
   END_STRUCT;
END_TYPE

TYPE "UDT_RP_MessageContFlush_v2"
VERSION : 0.1
   STRUCT
      xInitialized : Bool;   // The block is correctly initialized
      dNumOfMessage : DInt;   // Actual number of messages in buffer
      dMaxNumOfMessage : DInt;   // Maximum number of message in buffer
      rgtMessages : Array[0..12] of "UDT_RP_Message_v2";   // Array of messages
   END_STRUCT;
END_TYPE

TYPE "UDT_RP_Message_v2"
VERSION : 0.1
   STRUCT
      dCodeEvent : DInt;
      dtDateTime : Date_And_Time;
      strIdent : String[4];
      dEvent1 : DInt;
      dEvent2 : DInt;
      dEvent3 : DInt;
      dEvent4 : DInt;
      dEvent5 : DInt;
      dEvent6 : DInt;
      dEvent7 : DInt;
      dEvent8 : DInt;
      dEvent9 : DInt;
      dEvent10 : DInt;
   END_STRUCT;
END_TYPE

// folder: 09_Ribbon

TYPE "UDT_RibbonData"
   STRUCT
      dActualNumberGlassBreakMachine : DInt;   // Actual number of glass break machine
      dActualNumberGlassDataMachine : DInt;   // Actual number of glass data machine
      dActualNumberGlassThickMachine : DInt;   // Actual number of glass thickness machine
      rgtGlassBreak : Array[0.."DMAXGLASSBREAKMACHINE_IND"] of "UDT_RibbonData_GlassBreak";   // Glass break machine
      rgtGlassData : Array[0.."DMAXGLASSDATAMACHINE_IND"] of "UDT_RibbonData_GlassData";   // Glass data machine
      rgtGlassDataUpdate : Array[0.."DMAXGLASSDATAMACHINE_IND"] of Struct   // Structure where update the glass data status
         xUpdateRequest : Bool;   // Update request
         tData : "UDT_RibbonData_GlassData_SingleData";   // Actual data to use
      END_STRUCT;
      rgtGlassBreakUpdate : Array[0.."DMAXGLASSBREAKMACHINE_IND"] of Struct   // Structure where update the glass break status
         xUpdateRequest : Bool;   // Update request
         tData : "UDT_RibbonData_GlassBreak_SingleBreak";   // Actual data to use
      END_STRUCT;
      rgtGlassBreakRequest : Array[0.."DMAXGLASSBREAKREQUEST_IND"] of Struct   // Structure where get the break statuses
         IN_xRequestGlassBreak : Bool;   // Request glass break status at respective position
         IN_dDistanceSnaproll_cmm : DInt;   // Distance from snap roll [mm/100]
         IN_dUpstreamOffset_cmm : DInt;   // Upstream offset to anticipate the signal [mm/100]
         IN_dDownstreamOffset_cmm : DInt;   // Dowstream offset to retain the signal [mm/100]
         OUT_xDataReady : Bool;   // Data ready
         OUT_xGlassBreak : Bool;   // Glass break
      END_STRUCT;
      rgtGlassDataRequest : Array[0.."DMAXGLASSBREAKREQUEST_IND"] of Struct   // Structure where get the glass data statuses
         IN_xRequestGlassData : Bool;   // Request glass data at respective position
         IN_dDistanceSnaproll_cmm : DInt;   // Distance from snaproll [mm/100]
         IN_dSourceIndex : DInt;   // Index of the glass data source
         OUT_xDataReady : Bool;   // Data ready
         OUT_dGrossWidth_cmm : DInt;   // Actual gross width [mm/100]
         OUT_dNetWidth_cmm : DInt;   // Actual net width [mm/100]
         OUT_dGrossWander_cmm : DInt;   // Actual gross wander [mm/100]
         OUT_dNetWander_cmm : DInt;   // Actual net wander [mm/100]
      END_STRUCT;
   END_STRUCT;
END_TYPE

TYPE "UDT_RibbonData_GlassBreak"
   STRUCT
      dBufferHead : DInt := -1;   // Head of the glass data buffer
      dBufferTail : DInt := -1;   // Tail of the glass data buffer
      dLastInsertEncCount_cmm : DInt;   // Last insert encoder count [mm/100]
      dDistSnapRoll_cmm : DInt;   // Machine distance from snaproll [mm/100]
      rgtBuffer : Array[0.."DMAXGLASSBREAKSECTORS_IND"] of "UDT_RibbonData_GlassBreak_SingleBreak";   // Break buffer
      tLastDataBuffer : "UDT_RibbonData_GlassBreak_SingleBreak";   // Last break buffer
   END_STRUCT;
END_TYPE

TYPE "UDT_RibbonData_GlassBreak_SingleBreak"
   STRUCT
      xDataPresent : Bool;   // Item with valid data
      xUpdateDataBPSA : Bool;   // Update data on BPS A
      xUpdateDataBPSB : Bool;   // Update data on BPS B
      xGlassBreak : Bool;   // Glass break =1 Glass break in progress
      dEncoderValue_cmm : DInt;   // Actual encoder value [mm/100]
      rgxBreakMask : Array[0.."DMAXGLASSBREAKPHOTOCELL_IND"] of Bool;   // Activated photocell mask in this glass break
   END_STRUCT;
END_TYPE

TYPE "UDT_RibbonData_GlassData"
   STRUCT
      dBufferHead : DInt := -1;   // Head of the glass data buffer
      dBufferTail : DInt := -1;   // Tail of the glass data buffer
      dLastInsertEncCount_cmm : DInt;   // Last insert encoder count [mm/100]
      dDistSnapRoll_cmm : DInt;   // Machine distance from snaproll [mm/100]
      rgtBuffer : Array[0.."DMAXGLASSDATASECTORS_IND"] of "UDT_RibbonData_GlassData_SingleData";   // Glass data sectors
      tLastDataBuffer : "UDT_RibbonData_GlassData_SingleData";   // Last glass data buffer
   END_STRUCT;
END_TYPE

TYPE "UDT_RibbonData_GlassData_SingleData"
   STRUCT
      xDataPresent : Bool;   // Item with valid data
      xUpdateDataBPSA : Bool;   // Update data on BPS A
      xUpdateDataBPSB : Bool;   // Update data on BPS B
      dEncoderValue_cmm : DInt;   // Actual encoder value [mm/100]
      dGrossWidth_cmm : DInt;   // Actual gross width [mm/100]
      dNetWidth_cmm : DInt;   // Actual net width [mm/100]
      dGrossWander_cmm : DInt;   // Actual gross wander [mm/100]
      dNetWander_cmm : DInt;   // Actual net wander [mm/100]
   END_STRUCT;
END_TYPE

// folder: 10_Library

TYPE "UDT_IECTONTOFF_V1.00"
   STRUCT
      INTERNAL_dWaitingON_ms : DInt;   // Waiting ON timer
      INTERNAL_dRetainOFF_ms : DInt;   // Retain OFF timer
      INTERNAL_xLastSignalState : Bool;   // Last signal state
      INTERNAL_dLastTimeCount_ms : DInt;   // Last time count
      OUT_xDone : Bool;   // Timer done
   END_STRUCT;
END_TYPE

TYPE "UDT_IECTOFF_V1.00"
   STRUCT
      INTERNAL_dRetainOFF_ms : DInt;   // Retain OFF timer
      INTERNAL_xLastSignalState : Bool;   // Last signal state
      INTERNAL_dLastTimeCount_ms : DInt;   // Last time count
      OUT_xDone : Bool;   // Timer done
   END_STRUCT;
END_TYPE

TYPE "UDT_IECTON_V1.00"
   STRUCT
      INTERNAL_dWaitingON_ms : DInt;   // Waiting ON timer
      INTERNAL_xLastSignalState : Bool;   // Last signal state
      INTERNAL_dLastTimeCount_ms : DInt;   // Last time count
      OUT_xDone : Bool;   // Timer done
   END_STRUCT;
END_TYPE

// folder: 11_ConveyorMotorConfig

TYPE "UDT_MotorConfig"
   STRUCT
      iIOAddress_MM : Int;   // IO address motor module
      iPZD_MM : Int;   // Type of telegram(1=Open/closeLoop;111=Positioning)
      dMaxSpeed_rpm : DInt;   // Max Speed (set equal to StarterProject)[Rpm]
      rK_rpm_mmMin : Real;   // K Conversion From RPM to mm/min (value come from Drive)
      rK_mmMin_Rpm : Real;   // K Conversion From mm/min to Rpm (for Open Close Loop) value for Drive
      rMaxAcc : Real;   // Max Acceleration [Pos=m/s2, OpnLoop=S]
      rMaxDec : Real;   // Max Deceleration [Pos=m/s2, OpnLoop=S]
      rDec : Real;   // Deceleration [Pos=m/s2, OpnLoop=S]
      rAcc : Real;   // Acceleration [Pos=m/s2, OpnLoop=S]
      xModuleCorrect : Bool;   // Enable Module Correction
      xMDI_Continue : Bool;   // MDI
   END_STRUCT;
END_TYPE

// folder: 12_ProfinetDiagnostic

TYPE "TINFO_"
VERSION : 0.1
   STRUCT
      OB_start_info : Array[0..19] of Byte;
      W_20_STATION : Word;
      B22_slave_type : Byte;
      B23_interrupt_type : Byte;
      B24_origination : Byte;
      B25_diag_flag : Byte;
      W26_PN_ID : Word;
      W28_MFG_ID : Word;
      W30_INST_ID : Word;
      other_data : Array[1..70] of Byte;
   END_STRUCT;
END_TYPE

TYPE "AINFO_"
VERSION : 0.1
   STRUCT
      W0_block_type : Word;
      W2_block_length : Word;
      W4_version : Word;
      W6_interrupt_type : Word;
      D8_API : DWord;
      W12_comp_slot_num : Word;
      W14_submodule_slot_num : Word;
      D16_module_ID : DWord;
      D20_submodule_ID : DWord;
      W24_interrupt_specifer : Word;
      Add_W0_format_ID : Word;
      Add_W2_channel_num : Word;
      Add_B4_error_info : Byte;
      Add_B5_data_format : Byte;
      Add_W6_error_type : Word;
      extended_info : Array[34..1431] of Byte;
   END_STRUCT;
END_TYPE

TYPE "PN_Alarm"
VERSION : 0.1
   STRUCT
      word_allarme : Word;
      canale : Int;
   END_STRUCT;
END_TYPE

// folder: LGF/1 Date and timer operations

TYPE "LGF_typeGPS"
TITLE = LGF_typeGPS
// type for GPS Coordinates
   STRUCT
      latitude : "LGF_typeGPS_DMS";   // latitude child element
      longitude : "LGF_typeGPS_DMS";   // longitude child element
   END_STRUCT;
END_TYPE

TYPE "LGF_typeGPS_DD"
TITLE = LGF_typeGPS_DD
// type for GPS Coordinates in decimal degress
   STRUCT
      latitude : Real;   // latitude decimal degrees; North = positive; South = negative; [-90.0..90.0]
      longitude : Real;   // longitude decimal degrees; East=Positive; West = negative; [-180.0..180.0]
   END_STRUCT;
END_TYPE

TYPE "LGF_typeGPS_DMS"
TITLE = LGF_typeGPS_DMS
VERSION : 0.1
// type for GPS Coordinates for latitude OR longitude
   STRUCT
      dir : Char;   // Direction [N, S, E, W, n, s, e, w]
      deg : UInt;   // Degrees LAT [-89..+ 89]; LON [-179..+179]
      min : UInt;   // Minutes [0..+59]
      sec : UInt;   // Seconds [0..+59]
   END_STRUCT;
END_TYPE

// folder: (top level)

DATA_BLOCK "_debug"   // DB17
{ S7_Optimized_Access := 'TRUE' }
VERSION : 0.1
   VAR
      x : Bool;
      x1 : Bool;
      x2 : Bool;
      x3 : Bool;
      x4 : Bool;
      x5 : Bool;
      x6 : Bool;
      x7 : Bool;
      x8 : Bool;
      x9 : Bool;
      x10 : Bool;
   END_VAR
BEGIN
END_DATA_BLOCK

// folder: 03_Programs_Logics/MCC1200/03_CrossCut

DATA_BLOCK "DB_ExchangeDataModbus"   // DB63
{ S7_Optimized_Access := 'TRUE' }
VERSION : 0.1
   VAR
      Data : Array[0..39] of DInt;
      DataXcut : Array[0.."DMAXXHEADS_IND"] of Struct
         Data : Array[0..39] of DInt;
      END_STRUCT;
   END_VAR
BEGIN
END_DATA_BLOCK

DATA_BLOCK "DB_ExchangeDataModbusWrite"   // DB68
{ S7_Optimized_Access := 'TRUE' }
VERSION : 0.1
   VAR
      Data : Array[0..39] of DInt;
      DataXcut : Array[0.."DMAXXHEADS_IND"] of Struct
         Data : Array[0..39] of DInt;
      END_STRUCT;
   END_VAR
BEGIN
END_DATA_BLOCK

// folder: 03_Programs_Logics/MCC1200/15_ColdBackup

DATA_BLOCK "ExChangeParTxRx"   // DB187
{ S7_Optimized_Access := 'TRUE' }
VERSION : 0.1
   VAR
      tDataToSend : Struct
         dIndexParameter : DInt;   // Machine Index to Send
         dNByteBuffer : DInt;   // Number of byte in the buffer
         rgbBuffer : Array[0..500] of Byte;   // Buffer Parameter
      END_STRUCT;
      tDataRecived : Struct
         dIndexParameter : DInt;
         dNByteBuffer : DInt;   // Number of byte in the buffer
         rgbBuffer : Array[0..500] of Byte;   // FM152 - Temporary send buffer
      END_STRUCT;
      AUX_dIndexToSend : DInt;
      xRequestSend : Bool;
   END_VAR
BEGIN
END_DATA_BLOCK

DATA_BLOCK "FB_SwhitcTxRxColdBack_IDB"   // DB188
{ S7_Optimized_Access := 'TRUE' }
VERSION : 0.1
// stored: InstanceOfName FB_SwhitcTxRxColdBack_V1.00
"FB_SwhitcTxRxColdBack_V1.00"
BEGIN
END_DATA_BLOCK

// folder: 03_Programs_Logics/MCC1201/28_SpeedLehr

DATA_BLOCK "DB_AUX_Z200_SpeedLehr"   // DB80
{ S7_Optimized_Access := 'TRUE' }
VERSION : 0.1
   VAR
      dPulseEncoder1 : DInt;   // Pulse Encoder M200_BQ1.Encoder1
      dPulseEncoder2 : DInt;   // Pulse Encoder M200_BQ1.Encoder2
      dLastPulseEnc1 : DInt;   // Backup Pulse encoder 1
      dLastPulseEnc2 : DInt;   // Backup Pulse encoder 1
      dActualSpeedEncoder1 : DInt;   // Actual Speed [mm/min]
      dActualSpeedEncoder2 : DInt;   // Actual Speed [mm/min]
      tmON_LastBackupEnc1 : "UDT_IECTON_V1.00";   // Emergency OK timer / Last Backup encoder 1
      tmON_LastBackupEnc2 : "UDT_IECTON_V1.00";   // Emergency OK timer / Last Backup encoder 2
   END_VAR
BEGIN
END_DATA_BLOCK

// folder: 05_Reports

